// TIA Portal project "OpenLibraryExample" (V13) (continued)
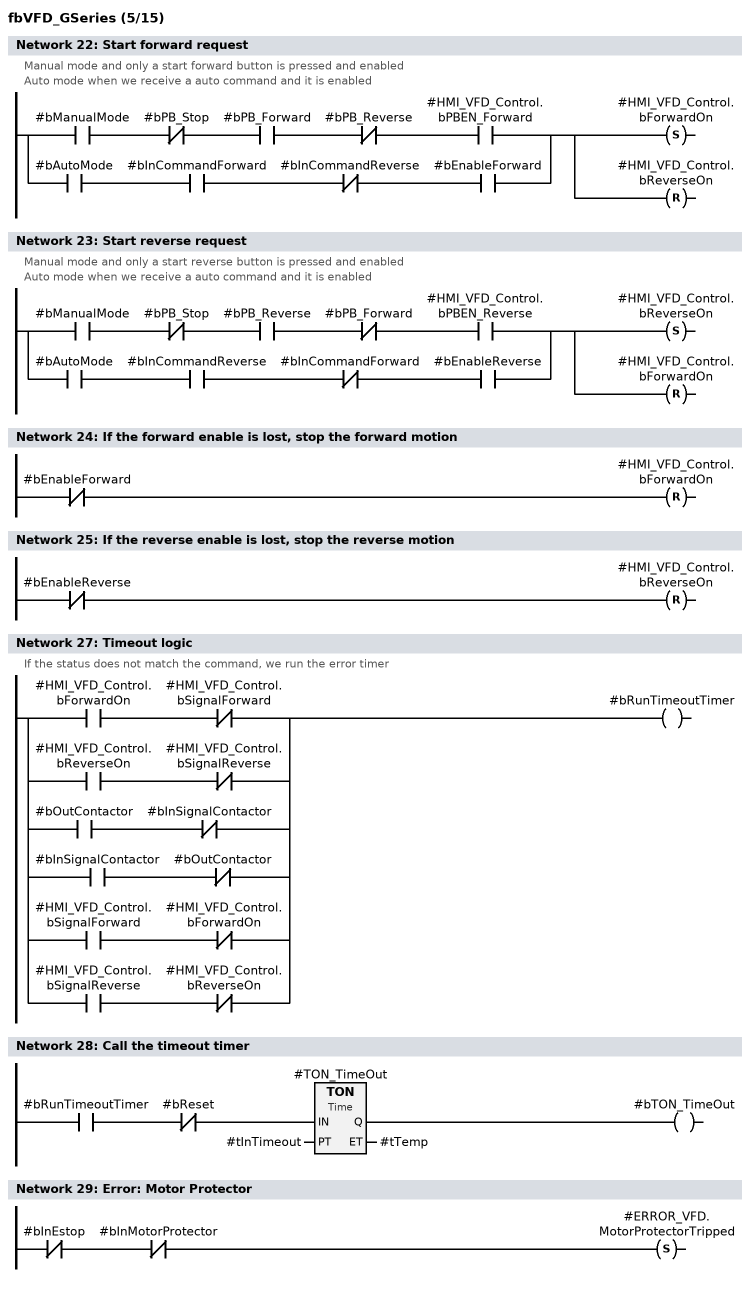
   RUNG wire#powerrail
      Contact( #bManualMode )
      I_Contact( #bPB_Stop )
      Contact( #bPB_Forward )
      I_Contact( #bPB_Reverse )
      Contact( #HMI_VFD_Control.bPBEN_Forward )
      wire#w1
      S_Coil( #HMI_VFD_Control.bForwardOn )
   END_RUNG
   RUNG wire#powerrail
      Contact( #bAutoMode )
      Contact( #bInCommandForward )
      I_Contact( #bInCommandReverse )
      Contact( #bEnableForward )
   END_RUNG wire#w1
   RUNG wire#w1
      R_Coil( #HMI_VFD_Control.bReverseOn )
   END_RUNG
   // the same network as SCL:
   IF (#bManualMode AND NOT #bPB_Stop AND #bPB_Forward AND NOT #bPB_Reverse AND #HMI_VFD_Control.bPBEN_Forward) OR (#bAutoMode AND #bInCommandForward AND NOT #bInCommandReverse AND #bEnableForward) THEN
       #HMI_VFD_Control.bForwardOn := TRUE;
       #HMI_VFD_Control.bReverseOn := FALSE;
   END_IF;
END_REGION

REGION Network 23: Start reverse request
   // Manual mode and only a start reverse button is pressed and enabled
   // Auto mode when we receive a auto command and it is enabled
   RUNG wire#powerrail
      Contact( #bManualMode )
      I_Contact( #bPB_Stop )
      Contact( #bPB_Reverse )
      I_Contact( #bPB_Forward )
      Contact( #HMI_VFD_Control.bPBEN_Reverse )
      wire#w1
      S_Coil( #HMI_VFD_Control.bReverseOn )
   END_RUNG
   RUNG wire#powerrail
      Contact( #bAutoMode )
      Contact( #bInCommandReverse )
      I_Contact( #bInCommandForward )
      Contact( #bEnableReverse )
   END_RUNG wire#w1
   RUNG wire#w1
      R_Coil( #HMI_VFD_Control.bForwardOn )
   END_RUNG
   // the same network as SCL:
   IF (#bManualMode AND NOT #bPB_Stop AND #bPB_Reverse AND NOT #bPB_Forward AND #HMI_VFD_Control.bPBEN_Reverse) OR (#bAutoMode AND #bInCommandReverse AND NOT #bInCommandForward AND #bEnableReverse) THEN
       #HMI_VFD_Control.bReverseOn := TRUE;
       #HMI_VFD_Control.bForwardOn := FALSE;
   END_IF;
END_REGION

REGION Network 24: If the forward enable is lost, stop the forward motion
   RUNG wire#powerrail
      I_Contact( #bEnableForward )
      R_Coil( #HMI_VFD_Control.bForwardOn )
   END_RUNG
   // the same network as SCL:
   IF NOT #bEnableForward THEN #HMI_VFD_Control.bForwardOn := FALSE; END_IF;
END_REGION

REGION Network 25: If the reverse enable is lost, stop the reverse motion
   RUNG wire#powerrail
      I_Contact( #bEnableReverse )
      R_Coil( #HMI_VFD_Control.bReverseOn )
   END_RUNG
   // the same network as SCL:
   IF NOT #bEnableReverse THEN #HMI_VFD_Control.bReverseOn := FALSE; END_IF;
END_REGION

REGION Network 26: --------------------------------------------------------- Errors ------------------------------------------------------------------
END_REGION

REGION Network 27: Timeout logic
   // If the status does not match the command, we run the error timer
   RUNG wire#powerrail
      Contact( #HMI_VFD_Control.bForwardOn )
      I_Contact( #HMI_VFD_Control.bSignalForward )
      wire#w1
      Coil( #bRunTimeoutTimer )
   END_RUNG
   RUNG wire#powerrail
      Contact( #HMI_VFD_Control.bReverseOn )
      I_Contact( #HMI_VFD_Control.bSignalReverse )
   END_RUNG wire#w1
   RUNG wire#powerrail
      Contact( #bOutContactor )
      I_Contact( #bInSignalContactor )
   END_RUNG wire#w1
   RUNG wire#powerrail
      Contact( #bInSignalContactor )
      I_Contact( #bOutContactor )
   END_RUNG wire#w1
   RUNG wire#powerrail
      Contact( #HMI_VFD_Control.bSignalForward )
      I_Contact( #HMI_VFD_Control.bForwardOn )
   END_RUNG wire#w1
   RUNG wire#powerrail
      Contact( #HMI_VFD_Control.bSignalReverse )
      I_Contact( #HMI_VFD_Control.bReverseOn )
   END_RUNG wire#w1
   // the same network as SCL:
   #bRunTimeoutTimer := (#HMI_VFD_Control.bForwardOn AND NOT #HMI_VFD_Control.bSignalForward) OR (#HMI_VFD_Control.bReverseOn AND NOT #HMI_VFD_Control.bSignalReverse) OR (#bOutContactor AND NOT #bInSignalContactor) OR (#bInSignalContactor AND NOT #bOutContactor) OR (#HMI_VFD_Control.bSignalForward AND NOT #HMI_VFD_Control.bForwardOn) OR (#HMI_VFD_Control.bSignalReverse AND NOT #HMI_VFD_Control.bReverseOn);
END_REGION

REGION Network 28: Call the timeout timer
   #TON_TimeOut.TON(IN := #bRunTimeoutTimer AND NOT #bReset, PT := #tInTimeout, ET => #tTemp);
   #bTON_TimeOut := #TON_TimeOut.Q;
END_REGION

REGION Network 29: Error: Motor Protector
   RUNG wire#powerrail
      I_Contact( #bInEstop )
      I_Contact( #bInMotorProtector )
      S_Coil( #ERROR_VFD.MotorProtectorTripped )
   END_RUNG
   // the same network as SCL:
   IF NOT #bInEstop AND NOT #bInMotorProtector THEN #ERROR_VFD.MotorProtectorTripped := TRUE; END_IF;
END_REGION

REGION Network 30: Error: Kill Switch/ local disconnect
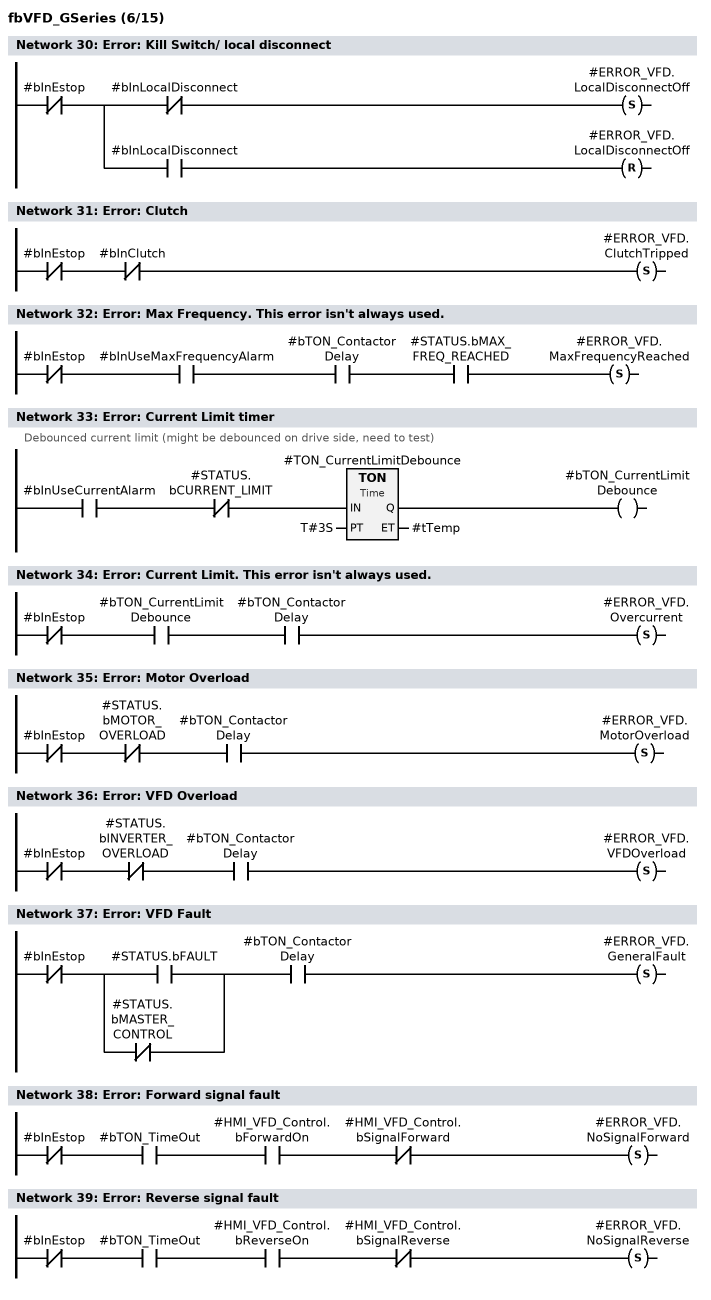
   RUNG wire#powerrail
      I_Contact( #bInEstop )
      wire#w1
      I_Contact( #bInLocalDisconnect )
      S_Coil( #ERROR_VFD.LocalDisconnectOff )
   END_RUNG
   RUNG wire#w1
      Contact( #bInLocalDisconnect )
      R_Coil( #ERROR_VFD.LocalDisconnectOff )
   END_RUNG
   // the same network as SCL:
   IF NOT #bInEstop AND NOT #bInLocalDisconnect THEN #ERROR_VFD.LocalDisconnectOff := TRUE; END_IF;
   IF NOT #bInEstop AND #bInLocalDisconnect THEN #ERROR_VFD.LocalDisconnectOff := FALSE; END_IF;
END_REGION

REGION Network 31: Error: Clutch
   RUNG wire#powerrail
      I_Contact( #bInEstop )
      I_Contact( #bInClutch )
      S_Coil( #ERROR_VFD.ClutchTripped )
   END_RUNG
   // the same network as SCL:
   IF NOT #bInEstop AND NOT #bInClutch THEN #ERROR_VFD.ClutchTripped := TRUE; END_IF;
END_REGION

REGION Network 32: Error: Max Frequency. This error isn't always used.
   RUNG wire#powerrail
      I_Contact( #bInEstop )
      Contact( #bInUseMaxFrequencyAlarm )
      Contact( #bTON_ContactorDelay )
      Contact( #STATUS.bMAX_FREQ_REACHED )
      S_Coil( #ERROR_VFD.MaxFrequencyReached )
   END_RUNG
   // the same network as SCL:
   IF NOT #bInEstop AND #bInUseMaxFrequencyAlarm AND #bTON_ContactorDelay AND #STATUS.bMAX_FREQ_REACHED THEN
       #ERROR_VFD.MaxFrequencyReached := TRUE;
   END_IF;
END_REGION

REGION Network 33: Error: Current Limit timer
   // Debounced current limit (might be debounced on drive side, need to test)
   #TON_CurrentLimitDebounce.TON(IN := #bInUseCurrentAlarm AND NOT #STATUS.bCURRENT_LIMIT,
                           PT := T#3S,
                           ET => #tTemp);
   #bTON_CurrentLimitDebounce := #TON_CurrentLimitDebounce.Q;
END_REGION

REGION Network 34: Error: Current Limit. This error isn't always used.
   RUNG wire#powerrail
      I_Contact( #bInEstop )
      Contact( #bTON_CurrentLimitDebounce )
      Contact( #bTON_ContactorDelay )
      S_Coil( #ERROR_VFD.Overcurrent )
   END_RUNG
   // the same network as SCL:
   IF NOT #bInEstop AND #bTON_CurrentLimitDebounce AND #bTON_ContactorDelay THEN
       #ERROR_VFD.Overcurrent := TRUE;
   END_IF;
END_REGION

REGION Network 35: Error: Motor Overload
   RUNG wire#powerrail
      I_Contact( #bInEstop )
      I_Contact( #STATUS.bMOTOR_OVERLOAD )
      Contact( #bTON_ContactorDelay )
      S_Coil( #ERROR_VFD.MotorOverload )
   END_RUNG
   // the same network as SCL:
   IF NOT #bInEstop AND NOT #STATUS.bMOTOR_OVERLOAD AND #bTON_ContactorDelay THEN
       #ERROR_VFD.MotorOverload := TRUE;
   END_IF;
END_REGION

REGION Network 36: Error: VFD Overload
   RUNG wire#powerrail
      I_Contact( #bInEstop )
      I_Contact( #STATUS.bINVERTER_OVERLOAD )
      Contact( #bTON_ContactorDelay )
      S_Coil( #ERROR_VFD.VFDOverload )
   END_RUNG
   // the same network as SCL:
   IF NOT #bInEstop AND NOT #STATUS.bINVERTER_OVERLOAD AND #bTON_ContactorDelay THEN
       #ERROR_VFD.VFDOverload := TRUE;
   END_IF;
END_REGION

REGION Network 37: Error: VFD Fault
   RUNG wire#powerrail
      I_Contact( #bInEstop )
      wire#w1
      Contact( #STATUS.bFAULT )
      wire#w2
      Contact( #bTON_ContactorDelay )
      S_Coil( #ERROR_VFD.GeneralFault )
   END_RUNG
   RUNG wire#w1
      I_Contact( #STATUS.bMASTER_CONTROL )
   END_RUNG wire#w2
   // the same network as SCL:
   IF NOT #bInEstop AND (#STATUS.bFAULT OR NOT #STATUS.bMASTER_CONTROL) AND #bTON_ContactorDelay THEN
       #ERROR_VFD.GeneralFault := TRUE;
   END_IF;
END_REGION

REGION Network 38: Error: Forward signal fault
   RUNG wire#powerrail
      I_Contact( #bInEstop )
      Contact( #bTON_TimeOut )
      Contact( #HMI_VFD_Control.bForwardOn )
      I_Contact( #HMI_VFD_Control.bSignalForward )
      S_Coil( #ERROR_VFD.NoSignalForward )
   END_RUNG
   // the same network as SCL:
   IF NOT #bInEstop AND #bTON_TimeOut AND #HMI_VFD_Control.bForwardOn AND NOT #HMI_VFD_Control.bSignalForward THEN
       #ERROR_VFD.NoSignalForward := TRUE;
   END_IF;
END_REGION

REGION Network 39: Error: Reverse signal fault
   RUNG wire#powerrail
      I_Contact( #bInEstop )
      Contact( #bTON_TimeOut )
      Contact( #HMI_VFD_Control.bReverseOn )
      I_Contact( #HMI_VFD_Control.bSignalReverse )
      S_Coil( #ERROR_VFD.NoSignalReverse )
   END_RUNG
   // the same network as SCL:
   IF NOT #bInEstop AND #bTON_TimeOut AND #HMI_VFD_Control.bReverseOn AND NOT #HMI_VFD_Control.bSignalReverse THEN
       #ERROR_VFD.NoSignalReverse := TRUE;
   END_IF;
END_REGION

REGION Network 40: Error: Motor contactor is not off
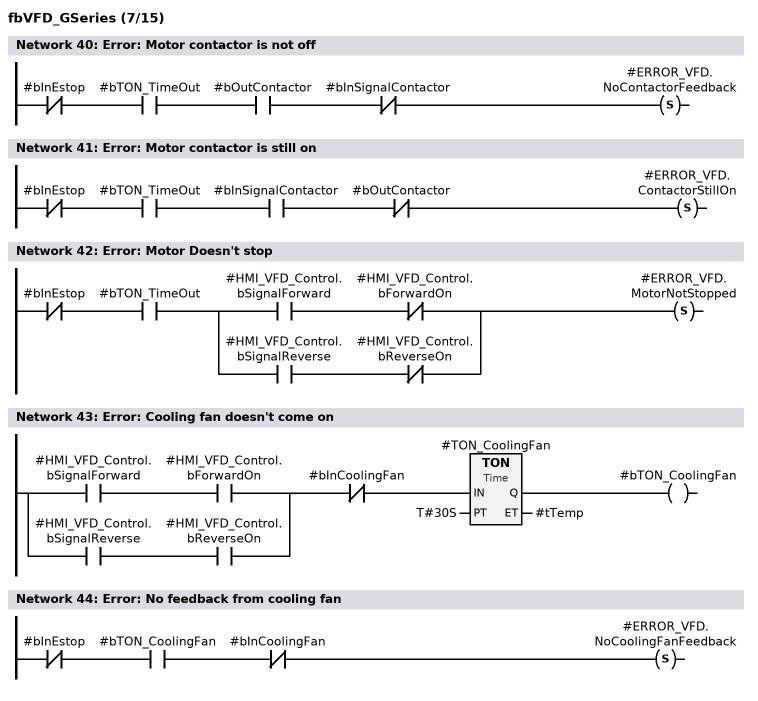
   RUNG wire#powerrail
      I_Contact( #bInEstop )
      Contact( #bTON_TimeOut )
      Contact( #bOutContactor )
      I_Contact( #bInSignalContactor )
      S_Coil( #ERROR_VFD.NoContactorFeedback )
   END_RUNG
   // the same network as SCL:
   IF NOT #bInEstop AND #bTON_TimeOut AND #bOutContactor AND NOT #bInSignalContactor THEN
       #ERROR_VFD.NoContactorFeedback := TRUE;
   END_IF;
END_REGION

REGION Network 41: Error: Motor contactor is still on
   RUNG wire#powerrail
      I_Contact( #bInEstop )
      Contact( #bTON_TimeOut )
      Contact( #bInSignalContactor )
      I_Contact( #bOutContactor )
      S_Coil( #ERROR_VFD.ContactorStillOn )
   END_RUNG
   // the same network as SCL:
   IF NOT #bInEstop AND #bTON_TimeOut AND #bInSignalContactor AND NOT #bOutContactor THEN
       #ERROR_VFD.ContactorStillOn := TRUE;
   END_IF;
END_REGION

REGION Network 42: Error: Motor Doesn't stop
   RUNG wire#powerrail
      I_Contact( #bInEstop )
      Contact( #bTON_TimeOut )
      wire#w1
      Contact( #HMI_VFD_Control.bSignalForward )
      I_Contact( #HMI_VFD_Control.bForwardOn )
      wire#w2
      S_Coil( #ERROR_VFD.MotorNotStopped )
   END_RUNG
   RUNG wire#w1
      Contact( #HMI_VFD_Control.bSignalReverse )
      I_Contact( #HMI_VFD_Control.bReverseOn )
   END_RUNG wire#w2
   // the same network as SCL:
   IF NOT #bInEstop AND #bTON_TimeOut AND ((#HMI_VFD_Control.bSignalForward AND NOT #HMI_VFD_Control.bForwardOn) OR (#HMI_VFD_Control.bSignalReverse AND NOT #HMI_VFD_Control.bReverseOn)) THEN
       #ERROR_VFD.MotorNotStopped := TRUE;
   END_IF;
END_REGION

REGION Network 43: Error: Cooling fan doesn't come on
   #TON_CoolingFan.TON(IN := ((#HMI_VFD_Control.bSignalForward AND #HMI_VFD_Control.bForwardOn) OR (#HMI_VFD_Control.bSignalReverse AND #HMI_VFD_Control.bReverseOn)) AND NOT #bInCoolingFan,
                       PT := T#30S,
                       ET => #tTemp);
   #bTON_CoolingFan := #TON_CoolingFan.Q;
END_REGION

REGION Network 44: Error: No feedback from cooling fan
   RUNG wire#powerrail
      I_Contact( #bInEstop )
      Contact( #bTON_CoolingFan )
      I_Contact( #bInCoolingFan )
      S_Coil( #ERROR_VFD.NoCoolingFanFeedback )
   END_RUNG
   // the same network as SCL:
   IF NOT #bInEstop AND #bTON_CoolingFan AND NOT #bInCoolingFan THEN
       #ERROR_VFD.NoCoolingFanFeedback := TRUE;
   END_IF;
END_REGION

REGION Network 45: Scroll errors on the HMI
   // Call the Error-Scroller which cyles through all possible errors and checks 
   // their state for display on the HMI
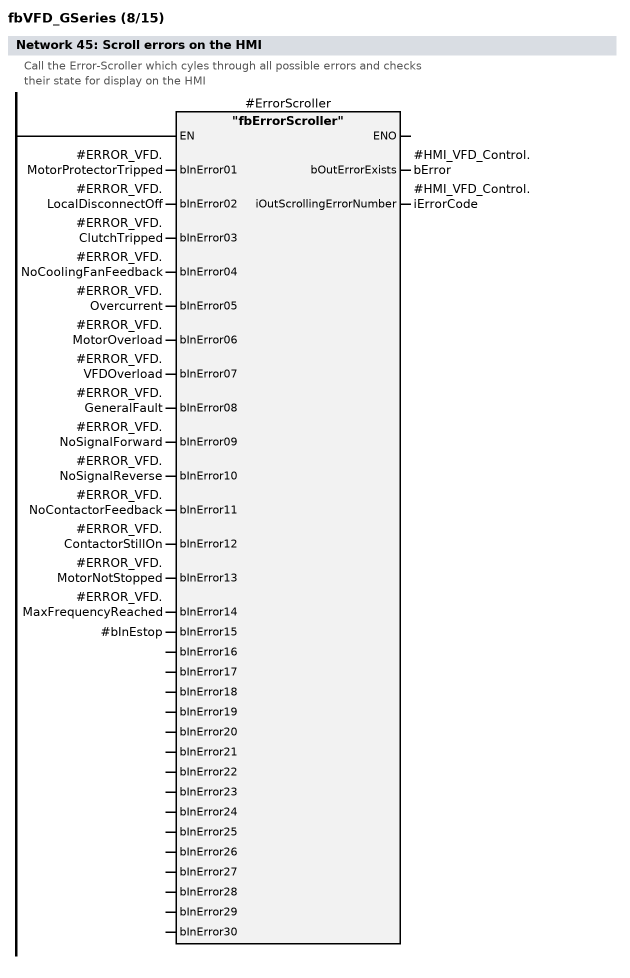
   RUNG wire#powerrail
      #ErrorScroller(bInError01 := #ERROR_VFD.MotorProtectorTripped, bInError02 := #ERROR_VFD.LocalDisconnectOff, bInError03 := #ERROR_VFD.ClutchTripped, bInError04 := #ERROR_VFD.NoCoolingFanFeedback, bInError05 := #ERROR_VFD.Overcurrent, bInError06 := #ERROR_VFD.MotorOverload, bInError07 := #ERROR_VFD.VFDOverload, bInError08 := #ERROR_VFD.GeneralFault, bInError09 := #ERROR_VFD.NoSignalForward, bInError10 := #ERROR_VFD.NoSignalReverse, bInError11 := #ERROR_VFD.NoContactorFeedback, bInError12 := #ERROR_VFD.ContactorStillOn, bInError13 := #ERROR_VFD.MotorNotStopped, bInError14 := #ERROR_VFD.MaxFrequencyReached, bInError15 := #bInEstop, bInError16 :=, bInError17 :=, bInError18 :=, bInError19 :=, bInError20 :=, bInError21 :=, bInError22 :=, bInError23 :=, bInError24 :=, bInError25 :=, bInError26 :=, bInError27 :=, bInError28 :=, bInError29 :=, bInError30 :=, bOutErrorExists => #HMI_VFD_Control.bError, iOutScrollingErrorNumber => #HMI_VFD_Control.iErrorCode)
   END_RUNG
   // the same network as SCL:
   #ErrorScroller(bInError01 := #ERROR_VFD.MotorProtectorTripped,   // "fbErrorScroller"
                  bInError02 := #ERROR_VFD.LocalDisconnectOff,
                  bInError03 := #ERROR_VFD.ClutchTripped,
                  bInError04 := #ERROR_VFD.NoCoolingFanFeedback,
                  bInError05 := #ERROR_VFD.Overcurrent,
                  bInError06 := #ERROR_VFD.MotorOverload,
                  bInError07 := #ERROR_VFD.VFDOverload,
                  bInError08 := #ERROR_VFD.GeneralFault,
                  bInError09 := #ERROR_VFD.NoSignalForward,
                  bInError10 := #ERROR_VFD.NoSignalReverse,
                  bInError11 := #ERROR_VFD.NoContactorFeedback,
                  bInError12 := #ERROR_VFD.ContactorStillOn,
                  bInError13 := #ERROR_VFD.MotorNotStopped,
                  bInError14 := #ERROR_VFD.MaxFrequencyReached,
                  bInError15 := #bInEstop,
                  bOutErrorExists => #HMI_VFD_Control.bError,
                  iOutScrollingErrorNumber => #HMI_VFD_Control.iErrorCode);
END_REGION

REGION Network 46: Set major fault bit
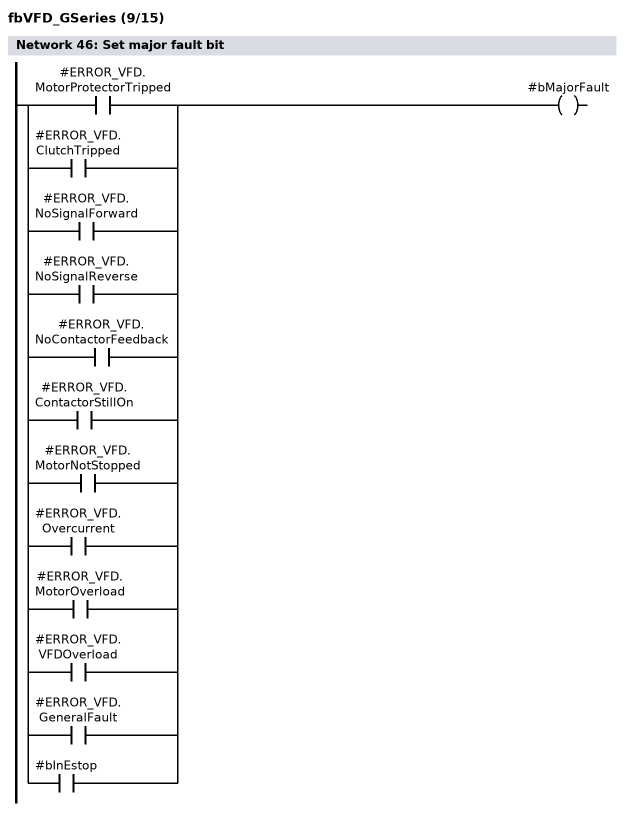
   RUNG wire#powerrail
      Contact( #ERROR_VFD.MotorProtectorTripped )
      wire#w1
      Coil( #bMajorFault )
   END_RUNG
   RUNG wire#powerrail
      Contact( #ERROR_VFD.ClutchTripped )
   END_RUNG wire#w1
   RUNG wire#powerrail
      Contact( #ERROR_VFD.NoSignalForward )
   END_RUNG wire#w1
   RUNG wire#powerrail
      Contact( #ERROR_VFD.NoSignalReverse )
   END_RUNG wire#w1
   RUNG wire#powerrail
      Contact( #ERROR_VFD.NoContactorFeedback )
   END_RUNG wire#w1
   RUNG wire#powerrail
      Contact( #ERROR_VFD.ContactorStillOn )
   END_RUNG wire#w1
   RUNG wire#powerrail
      Contact( #ERROR_VFD.MotorNotStopped )
   END_RUNG wire#w1
   RUNG wire#powerrail
      Contact( #ERROR_VFD.Overcurrent )
   END_RUNG wire#w1
   RUNG wire#powerrail
      Contact( #ERROR_VFD.MotorOverload )
   END_RUNG wire#w1
   RUNG wire#powerrail
      Contact( #ERROR_VFD.VFDOverload )
   END_RUNG wire#w1
   RUNG wire#powerrail
      Contact( #ERROR_VFD.GeneralFault )
   END_RUNG wire#w1
   RUNG wire#powerrail
      Contact( #bInEstop )
   END_RUNG wire#w1
   // the same network as SCL:
   #bMajorFault := #ERROR_VFD.MotorProtectorTripped OR #ERROR_VFD.ClutchTripped OR #ERROR_VFD.NoSignalForward OR #ERROR_VFD.NoSignalReverse OR #ERROR_VFD.NoContactorFeedback OR #ERROR_VFD.ContactorStillOn OR #ERROR_VFD.MotorNotStopped OR #ERROR_VFD.Overcurrent OR #ERROR_VFD.MotorOverload OR #ERROR_VFD.VFDOverload OR #ERROR_VFD.GeneralFault OR #bInEstop;
END_REGION

REGION Network 47: Set control bits based on major fault
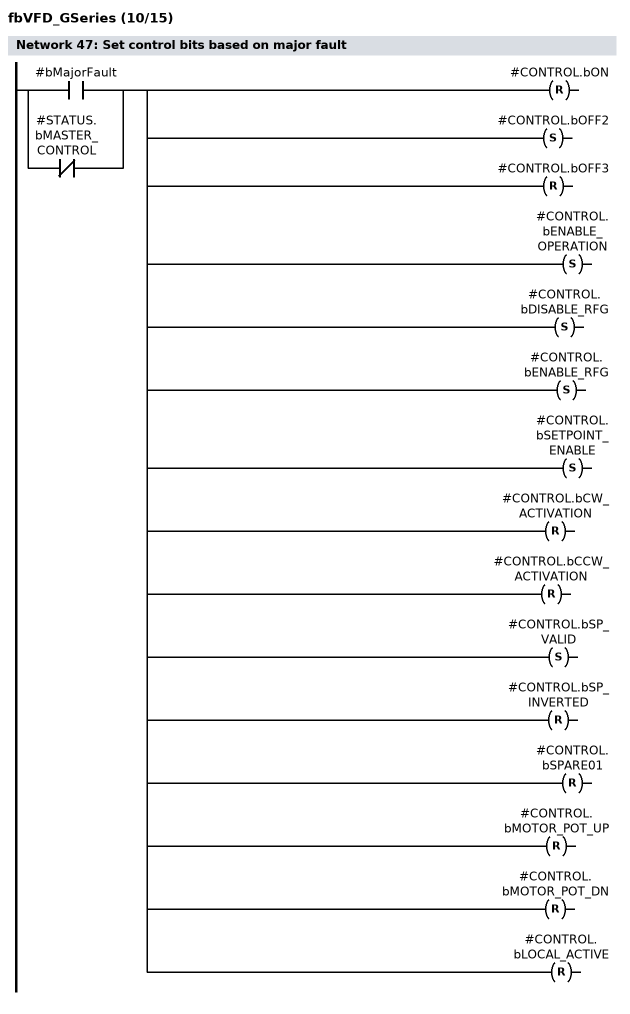
   RUNG wire#powerrail
      Contact( #bMajorFault )
      wire#w1
      R_Coil( #CONTROL.bON )
   END_RUNG
   RUNG wire#powerrail
      I_Contact( #STATUS.bMASTER_CONTROL )
   END_RUNG wire#w1
   RUNG wire#w1
      S_Coil( #CONTROL.bOFF2 )
   END_RUNG
   RUNG wire#w1
      R_Coil( #CONTROL.bOFF3 )
   END_RUNG
   RUNG wire#w1
      S_Coil( #CONTROL.bENABLE_OPERATION )
   END_RUNG
   RUNG wire#w1
      S_Coil( #CONTROL.bDISABLE_RFG )
   END_RUNG
   RUNG wire#w1
      S_Coil( #CONTROL.bENABLE_RFG )
   END_RUNG
   RUNG wire#w1
      S_Coil( #CONTROL.bSETPOINT_ENABLE )
   END_RUNG
   RUNG wire#w1
      R_Coil( #CONTROL.bCW_ACTIVATION )
   END_RUNG
   RUNG wire#w1
      R_Coil( #CONTROL.bCCW_ACTIVATION )
   END_RUNG
   RUNG wire#w1
      S_Coil( #CONTROL.bSP_VALID )
   END_RUNG
   RUNG wire#w1
      R_Coil( #CONTROL.bSP_INVERTED )
   END_RUNG
   RUNG wire#w1
      R_Coil( #CONTROL.bSPARE01 )
   END_RUNG
   RUNG wire#w1
      R_Coil( #CONTROL.bMOTOR_POT_UP )
   END_RUNG
   RUNG wire#w1
      R_Coil( #CONTROL.bMOTOR_POT_DN )
   END_RUNG
   RUNG wire#w1
      R_Coil( #CONTROL.bLOCAL_ACTIVE )
   END_RUNG
   // the same network as SCL:
   IF #bMajorFault OR NOT #STATUS.bMASTER_CONTROL THEN
       #CONTROL.bON := FALSE;
       #CONTROL.bOFF2 := TRUE;
       #CONTROL.bOFF3 := FALSE;
       #CONTROL.bENABLE_OPERATION := TRUE;
       #CONTROL.bDISABLE_RFG := TRUE;
       #CONTROL.bENABLE_RFG := TRUE;
       #CONTROL.bSETPOINT_ENABLE := TRUE;
       #CONTROL.bCW_ACTIVATION := FALSE;
       #CONTROL.bCCW_ACTIVATION := FALSE;
       #CONTROL.bSP_VALID := TRUE;
       #CONTROL.bSP_INVERTED := FALSE;
       #CONTROL.bSPARE01 := FALSE;
       #CONTROL.bMOTOR_POT_UP := FALSE;
       #CONTROL.bMOTOR_POT_DN := FALSE;
       #CONTROL.bLOCAL_ACTIVE := FALSE;
   END_IF;
END_REGION

REGION Network 48: Set control bits based on forward on command
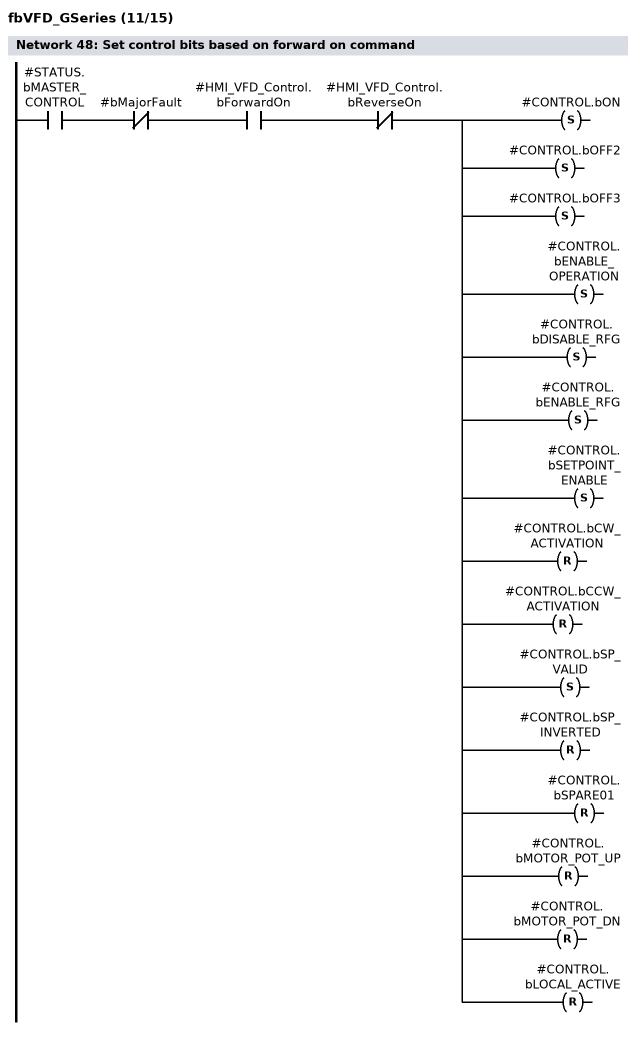
   RUNG wire#powerrail
      Contact( #STATUS.bMASTER_CONTROL )
      I_Contact( #bMajorFault )
      Contact( #HMI_VFD_Control.bForwardOn )
      I_Contact( #HMI_VFD_Control.bReverseOn )
      wire#w1
      S_Coil( #CONTROL.bON )
   END_RUNG
   RUNG wire#w1
      S_Coil( #CONTROL.bOFF2 )
   END_RUNG
   RUNG wire#w1
      S_Coil( #CONTROL.bOFF3 )
   END_RUNG
   RUNG wire#w1
      S_Coil( #CONTROL.bENABLE_OPERATION )
   END_RUNG
   RUNG wire#w1
      S_Coil( #CONTROL.bDISABLE_RFG )
   END_RUNG
   RUNG wire#w1
      S_Coil( #CONTROL.bENABLE_RFG )
   END_RUNG
   RUNG wire#w1
      S_Coil( #CONTROL.bSETPOINT_ENABLE )
   END_RUNG
   RUNG wire#w1
      R_Coil( #CONTROL.bCW_ACTIVATION )
   END_RUNG
   RUNG wire#w1
      R_Coil( #CONTROL.bCCW_ACTIVATION )
   END_RUNG
   RUNG wire#w1
      S_Coil( #CONTROL.bSP_VALID )
   END_RUNG
   RUNG wire#w1
      R_Coil( #CONTROL.bSP_INVERTED )
   END_RUNG
   RUNG wire#w1
      R_Coil( #CONTROL.bSPARE01 )
   END_RUNG
   RUNG wire#w1
      R_Coil( #CONTROL.bMOTOR_POT_UP )
   END_RUNG
   RUNG wire#w1
      R_Coil( #CONTROL.bMOTOR_POT_DN )
   END_RUNG
   RUNG wire#w1
      R_Coil( #CONTROL.bLOCAL_ACTIVE )
   END_RUNG
   // the same network as SCL:
   IF #STATUS.bMASTER_CONTROL AND NOT #bMajorFault AND #HMI_VFD_Control.bForwardOn AND NOT #HMI_VFD_Control.bReverseOn THEN
       #CONTROL.bON := TRUE;
       #CONTROL.bOFF2 := TRUE;
       #CONTROL.bOFF3 := TRUE;
       #CONTROL.bENABLE_OPERATION := TRUE;
       #CONTROL.bDISABLE_RFG := TRUE;
       #CONTROL.bENABLE_RFG := TRUE;
       #CONTROL.bSETPOINT_ENABLE := TRUE;
       #CONTROL.bCW_ACTIVATION := FALSE;
       #CONTROL.bCCW_ACTIVATION := FALSE;
       #CONTROL.bSP_VALID := TRUE;
       #CONTROL.bSP_INVERTED := FALSE;
       #CONTROL.bSPARE01 := FALSE;
       #CONTROL.bMOTOR_POT_UP := FALSE;
       #CONTROL.bMOTOR_POT_DN := FALSE;
       #CONTROL.bLOCAL_ACTIVE := FALSE;
   END_IF;
END_REGION

REGION Network 49: Set control bits based on Reverse on command
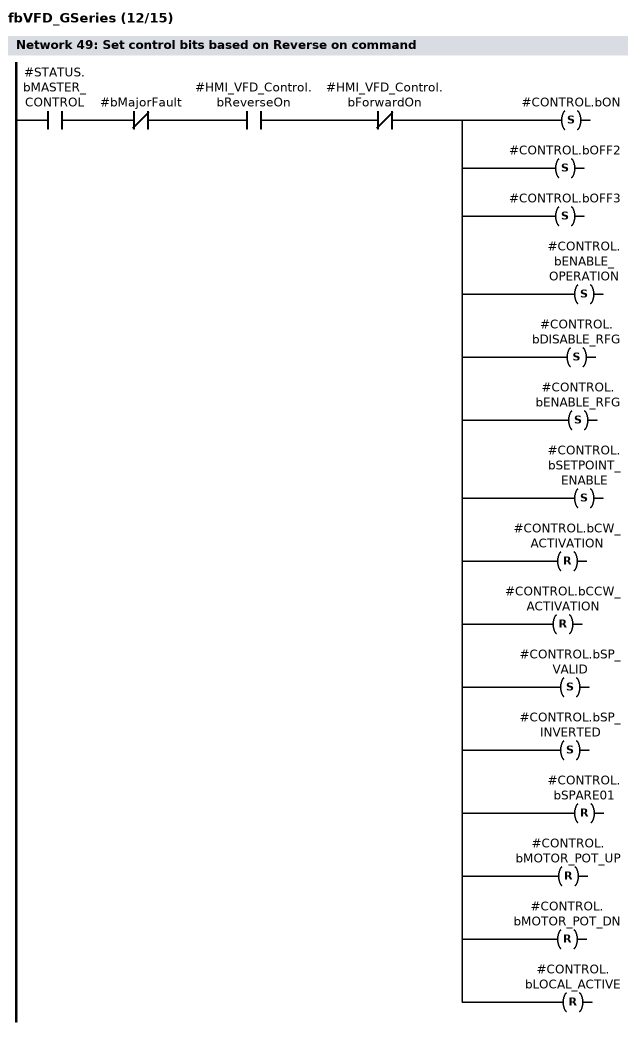
   RUNG wire#powerrail
      Contact( #STATUS.bMASTER_CONTROL )
      I_Contact( #bMajorFault )
      Contact( #HMI_VFD_Control.bReverseOn )
      I_Contact( #HMI_VFD_Control.bForwardOn )
      wire#w1
      S_Coil( #CONTROL.bON )
   END_RUNG
   RUNG wire#w1
      S_Coil( #CONTROL.bOFF2 )
   END_RUNG
   RUNG wire#w1
      S_Coil( #CONTROL.bOFF3 )
   END_RUNG
   RUNG wire#w1
      S_Coil( #CONTROL.bENABLE_OPERATION )
   END_RUNG
   RUNG wire#w1
      S_Coil( #CONTROL.bDISABLE_RFG )
   END_RUNG
   RUNG wire#w1
      S_Coil( #CONTROL.bENABLE_RFG )
   END_RUNG
   RUNG wire#w1
      S_Coil( #CONTROL.bSETPOINT_ENABLE )
   END_RUNG
   RUNG wire#w1
      R_Coil( #CONTROL.bCW_ACTIVATION )
   END_RUNG
   RUNG wire#w1
      R_Coil( #CONTROL.bCCW_ACTIVATION )
   END_RUNG
   RUNG wire#w1
      S_Coil( #CONTROL.bSP_VALID )
   END_RUNG
   RUNG wire#w1
      S_Coil( #CONTROL.bSP_INVERTED )
   END_RUNG
   RUNG wire#w1
      R_Coil( #CONTROL.bSPARE01 )
   END_RUNG
   RUNG wire#w1
      R_Coil( #CONTROL.bMOTOR_POT_UP )
   END_RUNG
   RUNG wire#w1
      R_Coil( #CONTROL.bMOTOR_POT_DN )
   END_RUNG
   RUNG wire#w1
      R_Coil( #CONTROL.bLOCAL_ACTIVE )
   END_RUNG
   // the same network as SCL:
   IF #STATUS.bMASTER_CONTROL AND NOT #bMajorFault AND #HMI_VFD_Control.bReverseOn AND NOT #HMI_VFD_Control.bForwardOn THEN
       #CONTROL.bON := TRUE;
       #CONTROL.bOFF2 := TRUE;
       #CONTROL.bOFF3 := TRUE;
       #CONTROL.bENABLE_OPERATION := TRUE;
       #CONTROL.bDISABLE_RFG := TRUE;
       #CONTROL.bENABLE_RFG := TRUE;
       #CONTROL.bSETPOINT_ENABLE := TRUE;
       #CONTROL.bCW_ACTIVATION := FALSE;
       #CONTROL.bCCW_ACTIVATION := FALSE;
       #CONTROL.bSP_VALID := TRUE;
       #CONTROL.bSP_INVERTED := TRUE;
       #CONTROL.bSPARE01 := FALSE;
       #CONTROL.bMOTOR_POT_UP := FALSE;
       #CONTROL.bMOTOR_POT_DN := FALSE;
       #CONTROL.bLOCAL_ACTIVE := FALSE;
   END_IF;
END_REGION

REGION Network 50: Set command bits when nothing is commanded, but no faults
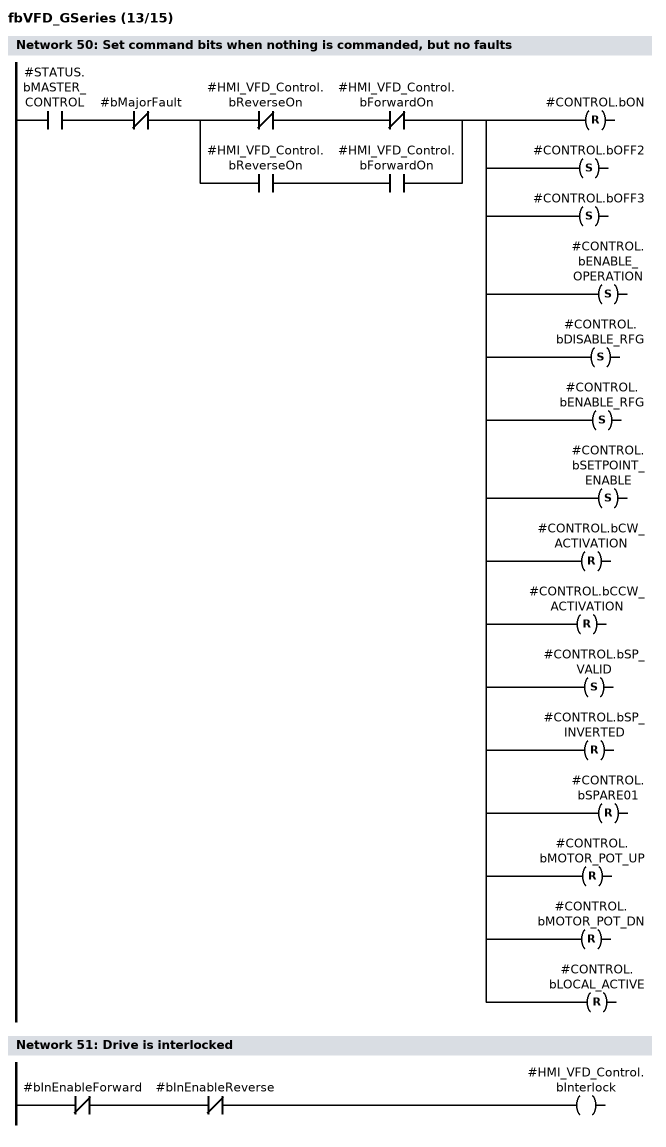
   RUNG wire#powerrail
      Contact( #STATUS.bMASTER_CONTROL )
      I_Contact( #bMajorFault )
      wire#w1
      I_Contact( #HMI_VFD_Control.bReverseOn )
      I_Contact( #HMI_VFD_Control.bForwardOn )
      wire#w2
      R_Coil( #CONTROL.bON )
   END_RUNG
   RUNG wire#w1
      Contact( #HMI_VFD_Control.bReverseOn )
      Contact( #HMI_VFD_Control.bForwardOn )
   END_RUNG wire#w2
   RUNG wire#w2
      S_Coil( #CONTROL.bOFF2 )
   END_RUNG
   RUNG wire#w2
      S_Coil( #CONTROL.bOFF3 )
   END_RUNG
   RUNG wire#w2
      S_Coil( #CONTROL.bENABLE_OPERATION )
   END_RUNG
   RUNG wire#w2
      S_Coil( #CONTROL.bDISABLE_RFG )
   END_RUNG
   RUNG wire#w2
      S_Coil( #CONTROL.bENABLE_RFG )
   END_RUNG
   RUNG wire#w2
      S_Coil( #CONTROL.bSETPOINT_ENABLE )
   END_RUNG
   RUNG wire#w2
      R_Coil( #CONTROL.bCW_ACTIVATION )
   END_RUNG
   RUNG wire#w2
      R_Coil( #CONTROL.bCCW_ACTIVATION )
   END_RUNG
   RUNG wire#w2
      S_Coil( #CONTROL.bSP_VALID )
   END_RUNG
   RUNG wire#w2
      R_Coil( #CONTROL.bSP_INVERTED )
   END_RUNG
   RUNG wire#w2
      R_Coil( #CONTROL.bSPARE01 )
   END_RUNG
   RUNG wire#w2
      R_Coil( #CONTROL.bMOTOR_POT_UP )
   END_RUNG
   RUNG wire#w2
      R_Coil( #CONTROL.bMOTOR_POT_DN )
   END_RUNG
   RUNG wire#w2
      R_Coil( #CONTROL.bLOCAL_ACTIVE )
   END_RUNG
   // the same network as SCL:
   IF #STATUS.bMASTER_CONTROL AND NOT #bMajorFault AND ((NOT #HMI_VFD_Control.bReverseOn AND NOT #HMI_VFD_Control.bForwardOn) OR (#HMI_VFD_Control.bReverseOn AND #HMI_VFD_Control.bForwardOn)) THEN
       #CONTROL.bON := FALSE;
       #CONTROL.bOFF2 := TRUE;
       #CONTROL.bOFF3 := TRUE;
       #CONTROL.bENABLE_OPERATION := TRUE;
       #CONTROL.bDISABLE_RFG := TRUE;
       #CONTROL.bENABLE_RFG := TRUE;
       #CONTROL.bSETPOINT_ENABLE := TRUE;
       #CONTROL.bCW_ACTIVATION := FALSE;
       #CONTROL.bCCW_ACTIVATION := FALSE;
       #CONTROL.bSP_VALID := TRUE;
       #CONTROL.bSP_INVERTED := FALSE;
       #CONTROL.bSPARE01 := FALSE;
       #CONTROL.bMOTOR_POT_UP := FALSE;
       #CONTROL.bMOTOR_POT_DN := FALSE;
       #CONTROL.bLOCAL_ACTIVE := FALSE;
   END_IF;
END_REGION

REGION Network 51: Drive is interlocked
   RUNG wire#powerrail
      I_Contact( #bInEnableForward )
      I_Contact( #bInEnableReverse )
      Coil( #HMI_VFD_Control.bInterlock )
   END_RUNG
   // the same network as SCL:
   #HMI_VFD_Control.bInterlock := NOT #bInEnableForward AND NOT #bInEnableReverse;
END_REGION

REGION Network 52: Set HMI status
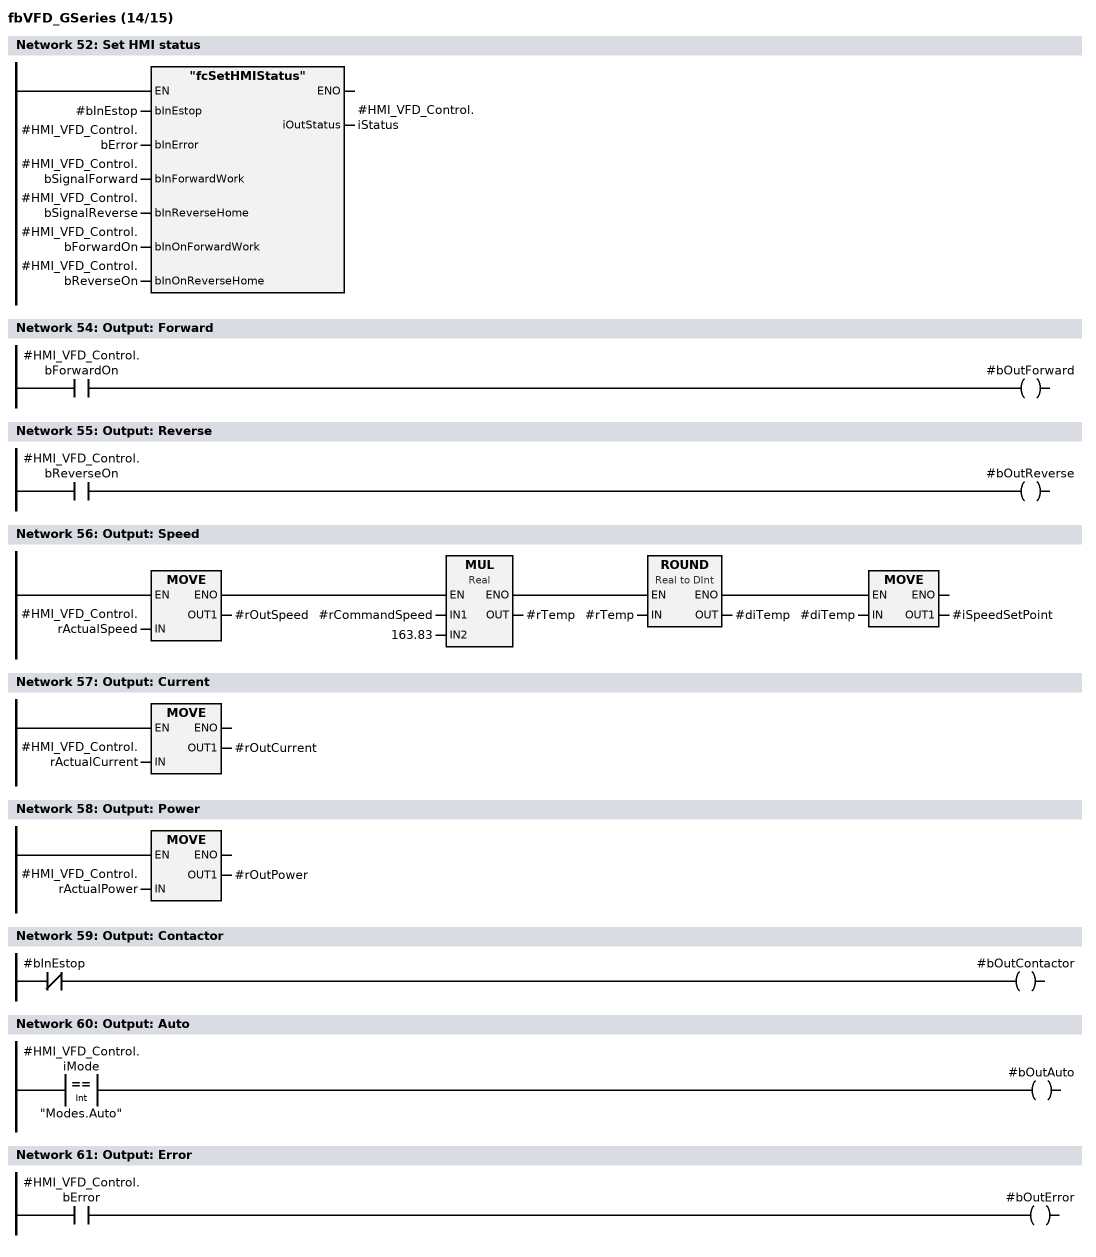
   RUNG wire#powerrail
      "fcSetHMIStatus"(bInEstop := #bInEstop, bInError := #HMI_VFD_Control.bError, bInForwardWork := #HMI_VFD_Control.bSignalForward, bInReverseHome := #HMI_VFD_Control.bSignalReverse, bInOnForwardWork := #HMI_VFD_Control.bForwardOn, bInOnReverseHome := #HMI_VFD_Control.bReverseOn, iOutStatus => #HMI_VFD_Control.iStatus)
   END_RUNG
   // the same network as SCL:
   "fcSetHMIStatus"(bInEstop := #bInEstop,
                    bInError := #HMI_VFD_Control.bError,
                    bInForwardWork := #HMI_VFD_Control.bSignalForward,
                    bInReverseHome := #HMI_VFD_Control.bSignalReverse,
                    bInOnForwardWork := #HMI_VFD_Control.bForwardOn,
                    bInOnReverseHome := #HMI_VFD_Control.bReverseOn,
                    iOutStatus => #HMI_VFD_Control.iStatus);
END_REGION

REGION Network 53: --------------------------------------------------------- Outputs ------------------------------------------------------------------
END_REGION

REGION Network 54: Output: Forward
   RUNG wire#powerrail
      Contact( #HMI_VFD_Control.bForwardOn )
      Coil( #bOutForward )
   END_RUNG
   // the same network as SCL:
   #bOutForward := #HMI_VFD_Control.bForwardOn;
END_REGION

REGION Network 55: Output: Reverse
   RUNG wire#powerrail
      Contact( #HMI_VFD_Control.bReverseOn )
      Coil( #bOutReverse )
   END_RUNG
   // the same network as SCL:
   #bOutReverse := #HMI_VFD_Control.bReverseOn;
END_REGION

REGION Network 56: Output: Speed
   RUNG wire#powerrail
      { S7_GenerateENO := "TRUE" } Move(in := #HMI_VFD_Control.rActualSpeed, out1 => #rOutSpeed)
      { S7_Templates := "SrcType := Real"; S7_GenerateENO := "TRUE" } Mul(in1 := #rCommandSpeed, in2 := 163.83, out => #rTemp)
      { S7_Templates := "[SrcType := Real, DestType := DInt]"; S7_GenerateENO := "TRUE" } Round(in := #rTemp, out => #diTemp)
      { S7_GenerateENO := "TRUE" } Move(in := #diTemp, out1 => #iSpeedSetPoint)
   END_RUNG
   // the same network as SCL:
   // ENO of a box is taken as its EN; it also drops when the box reports an error
   #rOutSpeed := #HMI_VFD_Control.rActualSpeed;
   #rTemp := #rCommandSpeed * 163.83;
   #diTemp := ROUND(#rTemp);
   #iSpeedSetPoint := #diTemp;
END_REGION

REGION Network 57: Output: Current
   RUNG wire#powerrail
      { S7_GenerateENO := "TRUE" } Move(in := #HMI_VFD_Control.rActualCurrent, out1 => #rOutCurrent)
   END_RUNG
   // the same network as SCL:
   #rOutCurrent := #HMI_VFD_Control.rActualCurrent;
END_REGION

REGION Network 58: Output: Power
   RUNG wire#powerrail
      { S7_GenerateENO := "TRUE" } Move(in := #HMI_VFD_Control.rActualPower, out1 => #rOutPower)
   END_RUNG
   // the same network as SCL:
   #rOutPower := #HMI_VFD_Control.rActualPower;
END_REGION

REGION Network 59: Output: Contactor
   RUNG wire#powerrail
      I_Contact( #bInEstop )
      Coil( #bOutContactor )
   END_RUNG
   // the same network as SCL:
   #bOutContactor := NOT #bInEstop;
END_REGION

REGION Network 60: Output: Auto
   RUNG wire#powerrail
      { S7_Templates := "SrcType := Int" } EQ_Contact(in1 := #HMI_VFD_Control.iMode, in2 := "Modes.Auto")
      Coil( #bOutAuto )
   END_RUNG
   // the same network as SCL:
   #bOutAuto := #HMI_VFD_Control.iMode = "Modes.Auto";
END_REGION

REGION Network 61: Output: Error
   RUNG wire#powerrail
      Contact( #HMI_VFD_Control.bError )
      Coil( #bOutError )
   END_RUNG
   // the same network as SCL:
   #bOutError := #HMI_VFD_Control.bError;
END_REGION

REGION Network 62: Output: Control Word
   // assemble control bits into control word
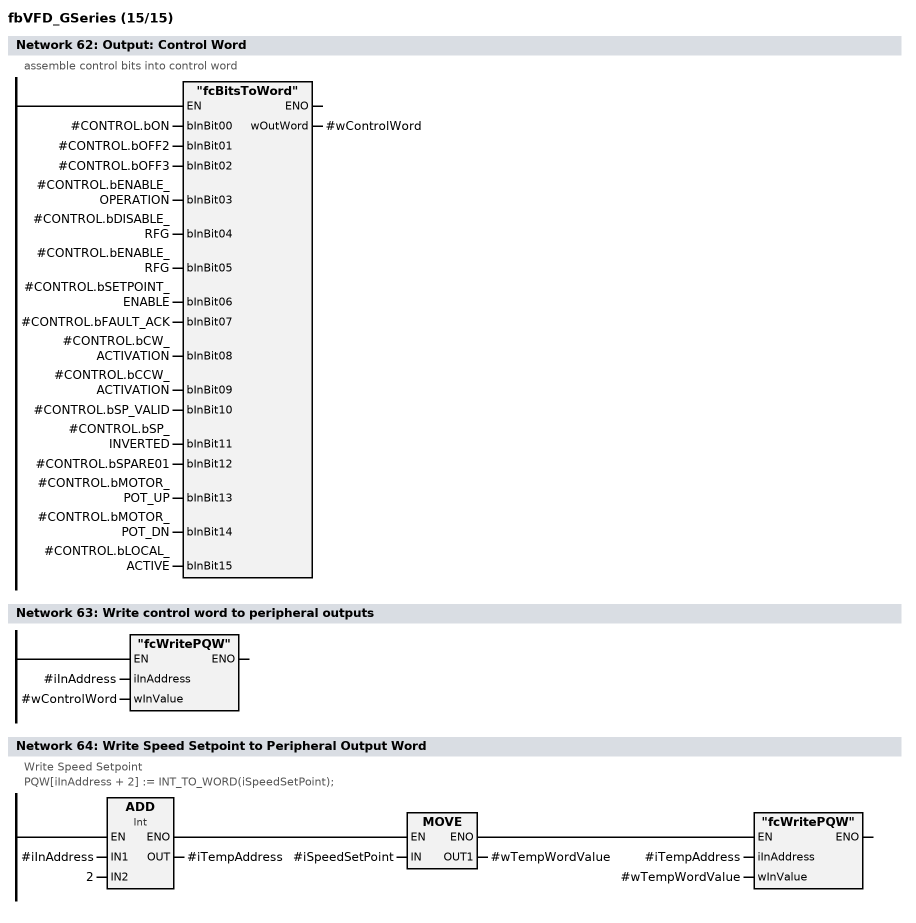
   RUNG wire#powerrail
      "fcBitsToWord"(bInBit00 := #CONTROL.bON, bInBit01 := #CONTROL.bOFF2, bInBit02 := #CONTROL.bOFF3, bInBit03 := #CONTROL.bENABLE_OPERATION, bInBit04 := #CONTROL.bDISABLE_RFG, bInBit05 := #CONTROL.bENABLE_RFG, bInBit06 := #CONTROL.bSETPOINT_ENABLE, bInBit07 := #CONTROL.bFAULT_ACK, bInBit08 := #CONTROL.bCW_ACTIVATION, bInBit09 := #CONTROL.bCCW_ACTIVATION, bInBit10 := #CONTROL.bSP_VALID, bInBit11 := #CONTROL.bSP_INVERTED, bInBit12 := #CONTROL.bSPARE01, bInBit13 := #CONTROL.bMOTOR_POT_UP, bInBit14 := #CONTROL.bMOTOR_POT_DN, bInBit15 := #CONTROL.bLOCAL_ACTIVE, wOutWord => #wControlWord)
   END_RUNG
   // the same network as SCL:
   "fcBitsToWord"(bInBit00 := #CONTROL.bON,
                  bInBit01 := #CONTROL.bOFF2,
                  bInBit02 := #CONTROL.bOFF3,
                  bInBit03 := #CONTROL.bENABLE_OPERATION,
                  bInBit04 := #CONTROL.bDISABLE_RFG,
                  bInBit05 := #CONTROL.bENABLE_RFG,
                  bInBit06 := #CONTROL.bSETPOINT_ENABLE,
                  bInBit07 := #CONTROL.bFAULT_ACK,
                  bInBit08 := #CONTROL.bCW_ACTIVATION,
                  bInBit09 := #CONTROL.bCCW_ACTIVATION,
                  bInBit10 := #CONTROL.bSP_VALID,
                  bInBit11 := #CONTROL.bSP_INVERTED,
                  bInBit12 := #CONTROL.bSPARE01,
                  bInBit13 := #CONTROL.bMOTOR_POT_UP,
                  bInBit14 := #CONTROL.bMOTOR_POT_DN,
                  bInBit15 := #CONTROL.bLOCAL_ACTIVE,
                  wOutWord => #wControlWord);
END_REGION

REGION Network 63: Write control word to peripheral outputs
   RUNG wire#powerrail
      "fcWritePQW"(iInAddress := #iInAddress, wInValue := #wControlWord)
   END_RUNG
   // the same network as SCL:
   "fcWritePQW"(iInAddress := #iInAddress, wInValue := #wControlWord);
END_REGION

REGION Network 64: Write Speed Setpoint to Peripheral Output Word
   // Write Speed Setpoint
   // PQW[iInAddress + 2] := INT_TO_WORD(iSpeedSetPoint);
   RUNG wire#powerrail
      { S7_Templates := "SrcType := Int"; S7_GenerateENO := "TRUE" } Add(in1 := #iInAddress, in2 := 2, out => #iTempAddress)
      { S7_GenerateENO := "TRUE" } Move(in := #iSpeedSetPoint, out1 => #wTempWordValue)
      "fcWritePQW"(iInAddress := #iTempAddress, wInValue := #wTempWordValue)
   END_RUNG
   // the same network as SCL:
   // ENO of a box is taken as its EN; it also drops when the box reports an error
   #iTempAddress := #iInAddress + 2;
   #wTempWordValue := #iSpeedSetPoint;
   "fcWritePQW"(iInAddress := #iTempAddress, wInValue := #wTempWordValue);
END_REGION
END_FUNCTION_BLOCK

FUNCTION_BLOCK "fbVFD_Analog"   // FB121, LAD
TITLE = Controls an analog VFD
{ S7_Optimized_Access := 'FALSE' }
VERSION : 0.1
   VAR_TEMP   // added for the SCL form of the ladder/FBD networks
      _w1 : Bool;
      _w2 : Bool;
      _w3 : Bool;
      _w4 : Bool;
   END_VAR
BEGIN

REGION Network 1: --------------------------------------------------------- Inputs ------------------------------------------------------------------
END_REGION

REGION Network 2: Read HMI input buttons
